// TIA Portal project "HEAT-1-CADIZ-V16" (V20) (continued)
REGION Network 5
   RUNG wire#powerrail
      "ToolChange_DB"(kukaCmdOpenCover := "kukaCmdOpenCover", kukaCmdCloseCover := "kukaCmdCloseCover", kukaCmdUnlockMps := "kukaCmdUnlockMps", kukaCmdSafeForChange := true, dockSensorToolInPosition := "dockSensorToolInPosition", dockSensorCoverClosed := "dockSensorCoverClosed", dockSensorCoverOpen := "dockSensorCoverOpen", robotSensorMpsUnlocked := "robotSensorMpsUnlocked", robotSensorMpsLocked := "robotSensorMpsLocked", robotSensorMpsCoupled := "robotSensorMpsCoupled", robotSensorMpsCtrlAirPressureOk := "robotSensorMpsCtrlAirPressureOk", resetFault :=, dockValveCoverOpenOn => "dockValveCoverOpenOn", dockValveCoverCloseOn => "dockValveCoverCloseOn", dockValveV2UnlockOn => "dockValveV2UnlockOn", kukaFeedbackDockCoverOpen => "kukaFeedbackDockCoverOpen", kukaFeedbackDockCoverClosed => "kukaFeedbackDockCoverClosed", kukaFeedbackRobotMpsUnlocked => "kukaFeedbackRobotMpsUnlocked", kukaFeedbackRobotMpsLocked => "kukaFeedbackRobotMpsLocked", kukaFeedbackRobotMpsCoupled => "kukaFeedbackRobotMpsCoupled", kukaFeedbackMpsCtrlAirPressureOk => "kukaFeedbackRobotMpsCtrlAirPressureOk", kukaFeedbackDockToolInPosition => "kukaFeedbackDockToolInPosition", diagStep =>, diagFault =>, diagFaultCode =>)
   END_RUNG
   // the same network as SCL:
   "ToolChange_DB"(kukaCmdOpenCover := "kukaCmdOpenCover",   // "ToolChange"
                   kukaCmdCloseCover := "kukaCmdCloseCover",
                   kukaCmdUnlockMps := "kukaCmdUnlockMps",
                   kukaCmdSafeForChange := true,
                   dockSensorToolInPosition := "dockSensorToolInPosition",
                   dockSensorCoverClosed := "dockSensorCoverClosed",
                   dockSensorCoverOpen := "dockSensorCoverOpen",
                   robotSensorMpsUnlocked := "robotSensorMpsUnlocked",
                   robotSensorMpsLocked := "robotSensorMpsLocked",
                   robotSensorMpsCoupled := "robotSensorMpsCoupled",
                   robotSensorMpsCtrlAirPressureOk := "robotSensorMpsCtrlAirPressureOk",
                   dockValveCoverOpenOn => "dockValveCoverOpenOn",
                   dockValveCoverCloseOn => "dockValveCoverCloseOn",
                   dockValveV2UnlockOn => "dockValveV2UnlockOn",
                   kukaFeedbackDockCoverOpen => "kukaFeedbackDockCoverOpen",
                   kukaFeedbackDockCoverClosed => "kukaFeedbackDockCoverClosed",
                   kukaFeedbackRobotMpsUnlocked => "kukaFeedbackRobotMpsUnlocked",
                   kukaFeedbackRobotMpsLocked => "kukaFeedbackRobotMpsLocked",
                   kukaFeedbackRobotMpsCoupled => "kukaFeedbackRobotMpsCoupled",
                   kukaFeedbackMpsCtrlAirPressureOk => "kukaFeedbackRobotMpsCtrlAirPressureOk",
                   kukaFeedbackDockToolInPosition => "kukaFeedbackDockToolInPosition");
END_REGION
END_FUNCTION_BLOCK

FUNCTION_BLOCK "SupervisorSeq"   // FB22, LAD
{ S7_Optimized_Access := 'TRUE' }
VERSION : 0.1
   VAR_INPUT
      T_Heartbeat : Time := T#1000ms;   // Periodo del heartbeat PLC
      T_IdCheck : Time := T#2000ms;   // Duración simulada de Identification (comprobaciones)
      enable : Bool;   // Habilita FB -> PLC.plc_ok
      QR_Ready : Bool;   // Hay un ID de carrito leído
      CarriageID : String;   // ID de carrito leído por QR
      TeachAtStart : Bool;   // Teaching (pág. 4): robot en punto de inicio de la siguiente trayectoria
      AtPerspex : Bool;   // PA check (Perspex) y Balancing (pág. 6): Robot posicionado en Perspex
      AtGainPos : Bool;   // Gain (pág. 7) -Robot posicionado para Gain
      AtTCGPos : Bool;   // TCG (pág. 8) — multiposición Robot en la posición TCG actual
      AtRefScanStart : Bool;   // Robot listo para Scan Ref
      AtInspScanStart : Bool;   // Robot listo para Scan Insp
      RefScanFinished : Bool;   // Trayectoria de referencia terminada (robot/UT)
      InspScanFinished : Bool;   // Trayectoria de inspección terminada (robot/UT)
      StartUSReady : Bool := TRUE;   // StartUS (pág. 5): end-effector y precondiciones listas -- True cuando “previous task done”
      MarkingDone : Bool;   // Pre-eval / marcado (pág. 13) -Resultado del marcado (true=OK)
      CmdStopUS : Bool;   // Orden local para Stop US
      CmdBreakUS : Bool;   // Pulso local Break US
      CmdUnbreakUS : Bool;   // Pulso local Unbreak US
   END_VAR
   VAR_OUTPUT
      ActiveStep : Int;   // Espejo local de PLC.step_plc
      AckSourceDbg : Int;   // Código de fuente de ACK (debug local)
      TCG_NextPosReq : Bool;   // PULSO 1 ciclo: mover a la SIGUIENTE posición TCG
      TCG_AdjustMode : Bool;   // LATCH: TRUE mientras estamos en “ajuste TCG”
   END_VAR
   VAR
      tHeartbeat : TON_TIME;
      tIdCheck : TON_TIME;
      hbGate : Bool;
      idCheckActive : Bool;
      prevStep : Int := -32768;
      firstScan : Bool;
      teachWasRunning : Bool;
      startUSWasRunning : Bool;
      elemWasRunning : Bool;
      balWasRunning : Bool;
      gainWasRunning : Bool;
      tcgWasInProgress : Bool;
      scanRefWasRunning : Bool;
      scanInspWasRunning : Bool;
      stopUSWasRunning : Bool;
      AckActive : Bool;   // ACK centralizado
      AckSource : Int;   // Qué petición estamos reconociendo
      evTCGNext : Bool;   // Eventos 1-ciclo que consume la máquina de estados
      evReqRefPart : Bool;
      evReqStopCycle : Bool;
      evReqTCGAdj : Bool;
      evReqVerif : Bool;
      evReqPreEval : Bool;
      evReqIdentState : Bool;
      carriageLatched : Bool;   // Otras memorias- para no reenviar ID cada ciclo
      mBreak : Bool;   // flanco Break US
      mUnbreak : Bool;   // flanco Unbreak US
      validScanParams : Bool;   // helper para scans
      waitingNextTCGPos : Bool;   // TRUE: esperar nueva posición antes de rearmar tcg_ready
   END_VAR
   VAR CONSTANT
      cSTEP_ID : Int := 1;   // // Pasos (según resumen del PDF, pág. 1)
      cSTEP_TEACH : Int := 2;
      cSTEP_STARTUS : Int := 3;
      cSTEP_PA_BAL : Int := 4;
      cSTEP_GAIN : Int := 5;
      cSTEP_TCG : Int := 6;
      cSTEP_SCAN_REF : Int := 7;
      cSTEP_SCAN_INSP : Int := 8;
      cSTEP_SCAN_REF_VERIF : Int := 9;
      cSTEP_PRE_EVAL : Int := 10;
      cACK_NONE : Int;   // // Fuentes de ACK (págs. 8, 11, 12)
      cACK_TCG_NEXT : Int := 1;
      cACK_REQ_REF : Int := 2;
      cACK_REQ_STOP : Int := 3;
      cACK_REQ_TCG_ADJ : Int := 4;
      cACK_REQ_VERIF : Int := 5;
      cACK_REQ_PRE_EVAL : Int := 6;
      cACK_REQ_IDENT_STATE : Int := 7;
   END_VAR
BEGIN

REGION Network 1 (SCL)
   // ------------------------------------------------------------------
   // 0) Servicios globales (Heartbeat, housekeeping) — vars generales (pág. 2)
   // ------------------------------------------------------------------
   "PlcStatus".plcOk := #enable;         // espejo de habilitación

   // Heartbeat PLC: toggle con TON (patrón de "compuerta")
   // hbGate se pone TRUE -> TON corre hasta PT -> tHeartbeat.Q = TRUE -> togglamos
   // y bajamos hbGate para reiniciar el ciclo.
   #tHeartbeat(IN := #hbGate,
               PT := #T_Heartbeat);
   IF NOT #hbGate THEN
       #hbGate := TRUE;
   ELSIF #tHeartbeat.Q THEN
       "PlcStatus".heartbeatPlc := NOT "PlcStatus".heartbeatPlc;
       #hbGate := FALSE;
   END_IF;

   // Normalizar paso y espejarlo a salida
   IF ("PlcStatus".stepPlc < #cSTEP_ID) OR ("PlcStatus".stepPlc > #cSTEP_PRE_EVAL) THEN
       "PlcStatus".stepPlc := #cSTEP_ID;
   END_IF;
   #ActiveStep := "PlcStatus".stepPlc;

   // firstScan: 1 ciclo al entrar en cada paso -> útil para resets seguros
   #firstScan := ("PlcStatus".stepPlc <> #prevStep);
   IF #firstScan THEN
       // Limpiamos cualquier "ready/start" que no deba arrastrarse al paso nuevo
       "PlcStatus".startUsReady := FALSE;
       "PlcStatus".stopUsReady := FALSE;
       "PlcStatus".paCheckReady := FALSE;
       "PlcStatus".gainReady := FALSE;
       "PlcStatus".tcgReady := FALSE;
       "PlcStatus".scanRefStart := FALSE;
       "PlcStatus".scanInspStart := FALSE;
       "PlcStatus".markRunning := FALSE;

       // reset de “había arrancado”
       #teachWasRunning := FALSE;
       #startUSWasRunning := FALSE;
       #elemWasRunning := FALSE;
       #balWasRunning := FALSE;
       #gainWasRunning := FALSE;
       #tcgWasInProgress := FALSE;
       #scanRefWasRunning := FALSE;
       #scanInspWasRunning := FALSE;

       // Señales generales de identificación
       "PlcStatus".idRunning := FALSE;

        //TCG: al entrar, exige confirmación de posición actual
       #waitingNextTCGPos := ("PlcStatus".stepPlc = #cSTEP_TCG) AND (NOT #AtTCGPos);
       // Salida auxiliar de ajuste TCG se limpia al cambiar de paso
       IF "PlcStatus".stepPlc <> #cSTEP_TCG THEN
           #TCG_AdjustMode := FALSE;
       END_IF;

       #prevStep := "PlcStatus".stepPlc;
   END_IF;

   // ------------------------------------------------------------------
   // [1] Gestor centralizado de ACK — TCG / Verif / PreEval / BackToID
   //     Idea: mientras una req_* esté a TRUE, PLC.acknowledge = TRUE.
   //     Cuando la req_* baja a FALSE, soltamos acknowledge y generamos
   //     un evento de 1 ciclo (evXXXX) para que el CASE tome decisiones.
   //     (ver págs. 8, 11, 12)
   // ------------------------------------------------------------------
   IF NOT #AckActive THEN
       // Tomamos la PRIMERA req_* que esté activa (prioridad de arriba a abajo)
       IF "SupervisorCmd".tcgNextStep THEN
           #AckActive := TRUE;
           #AckSource := #cACK_TCG_NEXT;
       ELSIF "SupervisorCmd".reqRefPart THEN
           #AckActive := TRUE;
           #AckSource := #cACK_REQ_REF;
       ELSIF "SupervisorCmd".reqStopCycle THEN
           #AckActive := TRUE;
           #AckSource := #cACK_REQ_STOP;
       ELSIF "SupervisorCmd".reqTcgAdj THEN
           #AckActive := TRUE;
           #AckSource := #cACK_REQ_TCG_ADJ;
       ELSIF "SupervisorCmd".reqVerif THEN
           #AckActive := TRUE;
           #AckSource := #cACK_REQ_VERIF;
       ELSIF "SupervisorCmd".reqPreEval THEN
           #AckActive := TRUE;
           #AckSource := #cACK_REQ_PRE_EVAL;
       ELSIF "SupervisorCmd".reqIdentificationState THEN
           #AckActive := TRUE;
           #AckSource := #cACK_REQ_IDENT_STATE;
       ELSE
           #AckSource := #cACK_NONE;
           #AckActive := FALSE;
       END_IF;
   END_IF;

   // Ejecutamos el reconocimiento según fuente
   CASE #AckSource OF
       #cACK_TCG_NEXT:
           "PlcStatus".acknowledge := TRUE;
           IF NOT "SupervisorCmd".tcgNextStep THEN
               // Fin del reconocimiento -> soltar y generar evento
               "PlcStatus".acknowledge := FALSE;
               #AckActive := FALSE;
               #AckSource := #cACK_NONE;
               #evTCGNext := TRUE;      // “pasar a siguiente pos” (p. 8)
           END_IF;

       #cACK_REQ_REF:
           "PlcStatus".acknowledge := TRUE;
           IF NOT "SupervisorCmd".reqRefPart THEN
               "PlcStatus".acknowledge := FALSE;
               #AckActive := FALSE;
               #AckSource := #cACK_NONE;
               #evReqRefPart := TRUE;// ir a Scan Ref (p. 8 → a)
           END_IF;

       #cACK_REQ_STOP:
           "PlcStatus".acknowledge := TRUE;
           IF NOT "SupervisorCmd".reqStopCycle THEN
               "PlcStatus".acknowledge := FALSE;
               #AckActive := FALSE;
               #AckSource := #cACK_NONE;
               #evReqStopCycle := TRUE; // cancelar ciclo (p. 8 → b)
           END_IF;

       #cACK_REQ_TCG_ADJ:
           "PlcStatus".acknowledge := TRUE;
           IF NOT "SupervisorCmd".reqTcgAdj THEN
               "PlcStatus".acknowledge := FALSE;
               #AckActive := FALSE;
               #AckSource := #cACK_NONE;
               #evReqTCGAdj := TRUE; // Seguir en TCG en modo ajuste (p. 8 → c)
           END_IF;

       #cACK_REQ_VERIF:
           "PlcStatus".acknowledge := TRUE;
           IF NOT "SupervisorCmd".reqVerif THEN
               "PlcStatus".acknowledge := FALSE;
               #AckActive := FALSE;
               #AckSource := #cACK_NONE;
               #evReqVerif := TRUE;   // Ir a verificación (p. 11)
           END_IF;

       #cACK_REQ_PRE_EVAL:
           "PlcStatus".acknowledge := TRUE;
           IF NOT "SupervisorCmd".reqPreEval THEN
               "PlcStatus".acknowledge := FALSE;
               #AckActive := FALSE;
               #AckSource := #cACK_NONE;
               #evReqPreEval := TRUE;  // Ir a Pre-eval (p. 12 → a)
           END_IF;

       #cACK_REQ_IDENT_STATE:
           "PlcStatus".acknowledge := TRUE;
           IF NOT "SupervisorCmd".reqIdentificationState THEN
               "PlcStatus".acknowledge := FALSE;
               #AckActive := FALSE;
               #AckSource := #cACK_NONE;
               #evReqIdentState := TRUE; //olver a Identification (p. 12 → b, p. 13)
           END_IF;

       ELSE
           "PlcStatus".acknowledge := FALSE;
   END_CASE;

   #AckSourceDbg := #AckSource;   // salida de diagnóstico local

   // ------------------------------------------------------------------
   // 2) MÁQUINA DE ESTADOS PRINCIPAL (CASE) — pasos del PDF
   // ------------------------------------------------------------------
   CASE "PlcStatus".stepPlc OF

           // ===============================================================
           // 1) IDENTIFICATION (pág. 3)
           // ===============================================================
       #cSTEP_ID:
           // --- Handshake de carriage ID ---
           // FÍSICO: lectura real de QR/PNs/params en HMI/Supervisor.
           // El PLC refleja ID leído y valida condiciones base (safety, agua, robot OK).
           // Supervisor.req_carriage_id = TRUE -> el PLC debe mandar:
           //   PLC.carriage_Id (string) y PLC.new_carriage_Id = TRUE
           // Mientras dure la petición. Al bajar la petición, el PLC
           // limpia new_carriage_Id y deja de enviar.
           // req_carriage_id: enviar ID nuevo UNA VEZ mientras Supervisor lo solicite
           IF "SupervisorCmd".reqCarriageId THEN
               IF #QR_Ready AND NOT #carriageLatched THEN
                   "PlcStatus".carriageId := #CarriageID; // escribimos el ID leído
                   "PlcStatus".newCarriageId := TRUE;     // “ID listo”
                   #carriageLatched := TRUE;              // evita rearmar en el mismo pulso
               END_IF;
           ELSE
               // fin del handshake
               "PlcStatus".newCarriageId := FALSE;
               #carriageLatched := FALSE;
           END_IF;

           // --- req_id -> identificación en curso ---
           // Cuando Supervisor pone req_id, el PLC indica id_running y,
           // tras un tiempo T_IdCheck, fija id_ok según condiciones globales.
           IF "SupervisorCmd".reqId AND NOT #idCheckActive THEN
               #idCheckActive := TRUE;
               "PlcStatus".idRunning := TRUE;
               "PlcStatus".idOk := FALSE;
               #tIdCheck(IN := TRUE,
                         PT := #T_IdCheck);  // arranca temporizador
           END_IF;

           IF #idCheckActive THEN
               #tIdCheck(IN := TRUE,
                         PT := #T_IdCheck);
               IF #tIdCheck.Q THEN
                   // Condiciones base (p. 2): enclavamientos / servicios / robot listo
                   "PlcStatus".idOk := ("PlcStatus".plcOk AND "SupervisorCmd".supervisorOk AND "PlcStatus".robotOk AND "PlcStatus".safetyOk
                   AND "PlcStatus".airOk AND "PlcStatus".inspWaterOk AND "PlcStatus".tankWaterOk);
                   "PlcStatus".idRunning := FALSE;
                   #idCheckActive := FALSE;
                   #tIdCheck(IN := FALSE,
                             PT := #T_IdCheck);

                   // Saltos según resultado y teach_req (pág. 3)
                   IF NOT "PlcStatus".idOk THEN
                       "PlcStatus".stepPlc := #cSTEP_ID; // cancelar ciclo / quedarse en identificación
                   ELSE
                       // Siguiente paso según teach_req (pág. 3)
                       IF "SupervisorCmd".teachReq THEN
                           "PlcStatus".stepPlc := #cSTEP_TEACH;
                       ELSE
                           "PlcStatus".stepPlc := #cSTEP_STARTUS;
                       END_IF;
                   END_IF;
               END_IF;
           ELSE
               // Aseguramos TON parado fuera del ciclo activo
               #tIdCheck(IN := FALSE,
                         PT := #T_IdCheck);
           END_IF;


           // ===============================================================
           // 2) TEACHING (pág. 4) — multi-PN: rearmar teach_ready por PN
           // FÍSICO: si la herramienta necesaria para teaching no está montada,
           // el KUKA cambia en Staübli al stand indicado (usa Supervisor.end-effector).
           // Luego, el KUKA se mueve al INICIO del PN siguiente y pone un bit de “en posición”.
           // Ese bit alimenta TeachAtStart=TRUE. Entonces EL PLC arma teach_ready (p. 4).
           // Repetir por cada PN mientras teach_app_running=TRUE.
           // ===============================================================
           (*  #cSTEP_TEACH:

            // Mientras la app de teaching esté abierta, debemos rearmar teach_ready
            // cada vez que el robot esté en el inicio del siguiente PN (TeachAtStart).
           IF "SupervisorCmd".teachAppRunning THEN
               // "Listo para enseñar" SOLO si NO está corriendo y robot en inicio PN              
               IF (NOT Supervisor.teach_running) AND #TeachAtStart THEN
                   "PlcStatus".teach_ready := TRUE; // // el láser/soft podrá iniciar teaching
               END_IF;

             // Al arrancar trayectoria de teaching -> soltamos ready
               IF Supervisor.teach_running THEN
                   PLC.teach_ready := FALSE;
                   #teachWasRunning := TRUE; // marcamos que empezó realmente
               END_IF;

                  // Al terminar una trayectoria (teach_running pasa a FALSE)
               IF (NOT Supervisor.teach_running) AND #teachWasRunning THEN
                   #teachWasRunning := FALSE; // fin de una trayectoria teaching
                    // Si siguen más PNs, se rearmará arriba (TeachAtStart=TRUE).
               END_IF;
           ELSE
                // Cierre de la app -> decidimos salto en base a teach_state (pág. 4)
               IF Supervisor.teach_state THEN
                   PLC.step_plc := #cSTEP_STARTUS;
               ELSE
                   PLC.step_plc := #cSTEP_ID;
               END_IF;
           END_IF;*)




           // ===============================================================
           // 3) START US (pág. 5) — armar cuando “previous task done”
           // FÍSICO: KUKA AUT EXT cambia (si hace falta) al efector de INSPECCIÓN
           // requerido (Supervisor.end-effector, p. 1). Cuando:
           //   - Herramienta correcta acoplada (Staübli OK),
           //   - servicios/enclavamientos OK (safety/air/water/tank),
           //   - robot en posición segura para inicializar el UT,
           // tu secuenciador pone StartUSReady=TRUE. El PLC arma start_us_ready.
           // Supervisor hace init UT (start_us_running/state_us). (p. 5)
           // ===============================================================
       #cSTEP_STARTUS:

           // Solo armamos start_us_ready si “previous task done” (StartUSReady)
           // y el Supervisor aún no ha arrancado.
           IF #StartUSReady AND NOT "SupervisorCmd".startUsRunning THEN
               "PlcStatus".startUsReady := TRUE; // → Supervisor puede iniciar
           END_IF;

           // Al comenzar la inicialización, soltamos el ready
           IF "SupervisorCmd".startUsRunning THEN
               "PlcStatus".startUsReady := FALSE;
               #startUSWasRunning := TRUE;
           END_IF;

           // Al finalizar la inicialización, Supervisor deja de correr y publica state_us
           IF (NOT "SupervisorCmd".startUsRunning) AND #startUSWasRunning THEN
               #startUSWasRunning := FALSE;
               IF NOT "SupervisorCmd".stateUs THEN
                   "PlcStatus".stepPlc := #cSTEP_ID; // fallo init US -> cancelar
               ELSE
                   IF "SupervisorCmd".paCheckReq THEN
                       "PlcStatus".stepPlc := #cSTEP_PA_BAL; // a) ir a PA-check (p. 5)
                   ELSE
                       "PlcStatus".stepPlc := #cSTEP_GAIN;   // b) ir a Gain (p. 5)
                   END_IF;
               END_IF;
           END_IF;

           // ===============================================================
           // 4) DEAD ELEMENT CHECK & BALANCING (pág. 6)
           //FÍSICO: KUKA va a la pieza Perspex de calibración y, cuando está en
           // posición estática, tu lógica pone AtPerspex=TRUE. El PLC arma
           // pa_check_ready y el Supervisor ejecuta elem_running/bal_running (p. 6).
           // ===============================================================
       #cSTEP_PA_BAL:

           // Dead elements en Perspex: el PLC pone pa_check_ready SOLO si
           // el robot ya está en la pieza Perspex y aún no corre elem_running
           IF #AtPerspex AND NOT "SupervisorCmd".elemRunning THEN
               "PlcStatus".paCheckReady := TRUE;
           END_IF;

           // Al iniciar la comprobación de dead elements soltamos ready
           IF "SupervisorCmd".elemRunning THEN
               "PlcStatus".paCheckReady := FALSE;
               #elemWasRunning := TRUE;
           END_IF;

           // Fin de dead elements -> miramos elem_state y encadenamos Balancing
           IF (NOT "SupervisorCmd".elemRunning) AND #elemWasRunning THEN
               #elemWasRunning := FALSE;
               IF NOT "SupervisorCmd".elemState THEN
                   "PlcStatus".stepPlc := #cSTEP_ID;
               ELSE
                   // Cascada a balancing (misma posición Perspex) (p. 6)
                   IF "SupervisorCmd".balRunning THEN
                       #balWasRunning := TRUE;
                   END_IF;

                   IF (NOT "SupervisorCmd".balRunning) AND #balWasRunning THEN
                       #balWasRunning := FALSE;
                       IF "SupervisorCmd".balState THEN
                           "PlcStatus".stepPlc := #cSTEP_GAIN;
                       ELSE
                           "PlcStatus".stepPlc := #cSTEP_ID;
                       END_IF;
                   END_IF;
               END_IF;
           END_IF;

           // ===============================================================
           // 5) GAIN ADJUSTMENT (pág. 7)
           // FÍSICO: KUKA se posiciona en la referencia para ganancia estática;
           // cuando está “en posición”, AtGainPos=TRUE. PLC arma gain_ready;
           // Supervisor ejecuta gain_running/gain_state y decide si ir a TCG (p. 7).
           // ===============================================================
       #cSTEP_GAIN:

           // Armamos gain_ready únicamente cuando el robot está en la posición
           // de ganancia y el supervisor todavía no corre la rutina de gain
           IF #AtGainPos AND NOT "SupervisorCmd".gainRunning THEN
               "PlcStatus".gainReady := TRUE;  // → Supervisor puede iniciar
           END_IF;

           IF "SupervisorCmd".gainRunning THEN
               "PlcStatus".gainReady := FALSE;
               #gainWasRunning := TRUE;
           END_IF;

           // Al terminar gain, ver resultado y decidir: TCG o Scan Ref
           IF (NOT "SupervisorCmd".gainRunning) AND #gainWasRunning THEN
               #gainWasRunning := FALSE;
               IF NOT "SupervisorCmd".gainState THEN
                   "PlcStatus".stepPlc := #cSTEP_ID;
               ELSE
                   IF "SupervisorCmd".tcgReq THEN
                       "PlcStatus".stepPlc := #cSTEP_TCG;
                   ELSE
                       "PlcStatus".stepPlc := #cSTEP_SCAN_REF;
                   END_IF;
               END_IF;
           END_IF;

           // ===============================================================
           // (6) TCG CHECK / ADJUSTMENT — pág. 8 (multiposición)
           // FÍSICO: KUKA recorre varias posiciones TCG. Para cada posición:
           //   - Cuando el robot está en la POSICIÓN TCG ACTUAL (estático),
           //     tu lógica pone AtTCGPos=TRUE → PLC arma tcg_ready (p. 8).
           //   - Supervisor pone tcg_in_progress=TRUE mientras mide.
           //   - Al pulsar “Next” en Supervisor (tcg_next_step=TRUE), el ACK manager
           //     emite TCG_NextPosReq (pulso) para que MUEVAS el robot a la SIGUIENTE
           //     posición; el FB bloquea el rearme (waitingNextTCGPos=TRUE) hasta que
           //     AtTCGPos vuelva a TRUE en la nueva posición (antirrebote).
           //   - Final: según req_ref_part / req_stop_cycle / req_tcg_adj (p. 8).
           // ===============================================================
       #cSTEP_TCG:

           // Confirmación de nueva posición alcanzada
           IF #waitingNextTCGPos AND #AtTCGPos THEN
               #waitingNextTCGPos := FALSE;     // nueva pos OK → se podrá rearmar ready
           END_IF;

           // Armado defensivo: tcg_ready SOLO si no hay progreso y no esperamos pos
           IF (NOT "SupervisorCmd".tcgInProgress) AND (NOT #waitingNextTCGPos) THEN
               "PlcStatus".tcgReady := TRUE;          // listo para medir en esta pos (p. 8)
           END_IF;

           IF "SupervisorCmd".tcgInProgress THEN
               "PlcStatus".tcgReady := FALSE;
               #tcgWasInProgress := TRUE;
           END_IF;

           // “Next” → mueve a la SIGUIENTE pos (tu secuenciador KUKA)
           IF #evTCGNext THEN
               #TCG_NextPosReq := TRUE;      // pulso 1 ciclo hacia tu lógica
               #waitingNextTCGPos := TRUE;      // bloquea ready hasta nueva posición
           END_IF;

           // “Ajuste TCG”
           IF #evReqTCGAdj THEN
               #TCG_AdjustMode := TRUE;        // permanecer en step 6 hasta validar
           END_IF;

           // Validación de TCG
           IF #evReqRefPart THEN
               #TCG_AdjustMode := FALSE;
               "PlcStatus".stepPlc := #cSTEP_SCAN_REF; // TCG OK → Scan Ref (p. 8)
           ELSIF #evReqStopCycle THEN
               #TCG_AdjustMode := FALSE;
               "PlcStatus".stepPlc := #cSTEP_ID;       // cancelar (p. 8)
           END_IF;



           // ===============================================================
           // (7) SCAN REFERENCE ACQUISITION — pág. 10
           // FÍSICO: KUKA carga PN/frame y se coloca en el punto de INICIO de
           // la trayectoria de referencia. Tu lógica pone AtRefScanStart=TRUE cuando
           // está en posición. El PLC solo arma scan_ref_start si además los
           // parámetros mínimos (id_scan, x_size, y_size) están válidos (p. 10).
           // ===============================================================
       #cSTEP_SCAN_REF:

           // Validación mínima de parámetros: hay PN/Frame y tamaños > 0.
           // (El PDF indica que el PLC envía id_scan, point_origin, x_size, y_size).
           #validScanParams := (LEN("PlcStatus".idScan) > 0) AND ("PlcStatus".xSize > 0.0) AND ("PlcStatus".ySize > 0.0);

           // "Robot ready" solo si parámetros OK, robot en inicio y aún no corre
           IF #AtRefScanStart AND #validScanParams AND NOT "SupervisorCmd".scanRefRunning THEN
               "PlcStatus".scanRefStart := TRUE;     // Supervisor cargará/validará y pondrá scan_ref_running
           END_IF;

           // En ejecución: opcionalmente bajar start al terminar la trayectoria
           IF "SupervisorCmd".scanRefRunning THEN
               #scanRefWasRunning := TRUE;
               IF #RefScanFinished THEN
                   "PlcStatus".scanRefStart := FALSE; // indica “fin de movimiento -> guardar”
               END_IF;
           END_IF;

           // Al terminar guardado, Supervisor baja running y publica scan_ref_state
           IF (NOT "SupervisorCmd".scanRefRunning) AND #scanRefWasRunning THEN
               #scanRefWasRunning := FALSE;
               "PlcStatus".scanRefStart := FALSE;
               IF NOT "SupervisorCmd".scanRefState THEN
                   "PlcStatus".stepPlc := #cSTEP_ID;   // error durante ref -> cancelar
               ELSE
                   "PlcStatus".stepPlc := #cSTEP_SCAN_INSP;
               END_IF;
           END_IF;

           // ===============================================================
           // (8) SCAN INSPECTION — pág. 11
           // FÍSICO: KUKA se coloca en INICIO de la(s) trayectoria(s) de inspección
           // (AtInspScanStart=TRUE). El PLC arma scan_insp_start solo si parámetros
           // válidos. Supervisor corre/guarda y luego pide verificación (req_verif) (p. 11).
           // ===============================================================
       #cSTEP_SCAN_INSP:

           // Validación mínima de parámetros: hay PN/Frame y tamaños > 0.
           // (El PDF indica que el PLC envía id_scan, point_origin, x_size, y_size).
           #validScanParams := (LEN("PlcStatus".idScan) > 0) AND ("PlcStatus".xSize > 0.0) AND ("PlcStatus".ySize > 0.0);

           // "Robot ready" solo si parámetros OK, robot en inicio y aún no corre
           IF #AtInspScanStart AND #validScanParams AND NOT "SupervisorCmd".scanInsprunning THEN
               "PlcStatus".scanInspStart := TRUE;    // Supervisor cargará y arrancará
           END_IF;

           // En ejecución: opcionalmente bajar start al terminar la trayectoria
           IF "SupervisorCmd".scanInsprunning THEN
               #scanInspWasRunning := TRUE;
               IF #InspScanFinished THEN
                   "PlcStatus".scanInspStart := FALSE; // fin de movimiento -> guardar
               END_IF;
           END_IF;

           // Al terminar guardado, Supervisor baja running y publica scan_ref_state
           IF (NOT "SupervisorCmd".scanInsprunning) AND #scanInspWasRunning THEN
               #scanInspWasRunning := FALSE;
               "PlcStatus".scanInspStart := FALSE;

               IF NOT "SupervisorCmd".scanInspState THEN
                   "PlcStatus".stepPlc := #cSTEP_ID;   // error -> cancelar
               ELSE
                   // Ir a verificación cuando el ACK manager confirme req_verif
                   IF #evReqVerif THEN
                       "PlcStatus".stepPlc := #cSTEP_SCAN_REF_VERIF;
                   END_IF;
               END_IF;
           END_IF;


           // ===============================================================
           // (9) SCAN REFERENCE VERIFICATION — pág. 12
           // FÍSICO: KUKA vuelve al INICIO de la trayectoria de verificación de ref.
           // (AtRefScanStart=TRUE). Igual patrón de parámetros/ready/running/state (p. 12).
           // Fin: Supervisor decide Pre‑eval (req_pre_eval) o nuevo ciclo (req_identification_state).
           // ===============================================================
       #cSTEP_SCAN_REF_VERIF:

           #validScanParams := (LEN("PlcStatus".idScan) > 0) AND ("PlcStatus".xSize > 0.0) AND ("PlcStatus".ySize > 0.0);

           IF #AtRefScanStart AND #validScanParams AND NOT "SupervisorCmd".scanRefRunning THEN
               "PlcStatus".scanRefStart := TRUE;     // Robot listo para verificación de ref
           END_IF;

           IF "SupervisorCmd".scanRefRunning THEN
               #scanRefWasRunning := TRUE;
           END_IF;

           IF (NOT "SupervisorCmd".scanRefRunning) AND #scanRefWasRunning THEN
               #scanRefWasRunning := FALSE;
               "PlcStatus".scanRefStart := FALSE;

               IF NOT "SupervisorCmd".scanRefState THEN
                   "PlcStatus".stepPlc := #cSTEP_ID;
               ELSE
                   // a) Pre‑eval   b) Volver a Identification
                   IF #evReqPreEval THEN
                       "PlcStatus".stepPlc := #cSTEP_PRE_EVAL;
                   ELSIF #evReqIdentState THEN
                       "PlcStatus".stepPlc := #cSTEP_ID;
                   END_IF;
               END_IF;
           END_IF;

           // ===============================================================
           // (10) PRE‑EVALUATION / MARKING — pág. 13
           // FÍSICO: si la herramienta de marcado no está montada, el KUKA cambia
           // en Staübli al stand de “marking” según requiera el proceso; tras estar
           // listo se puede marcar (Supervisor.req_mark). El resultado físico del
           // marcado tu lógica lo refleja en MarkingDone=TRUE/FALSE (p. 13).
           // También se puede arrancar un nuevo ciclo (req_identification_state).
           // ===============================================================
       #cSTEP_PRE_EVAL:

           // b) Volver a inicio (nuevo ciclo)
           IF #evReqIdentState THEN
               "PlcStatus".stepPlc := #cSTEP_ID;
           END_IF;

           // a) Marcado: si Supervisor.req_mark, ejecutamos el ciclo simple:
           //   - mark_running TRUE durante la acción
           //   - mark_state según resultado físico (MarkingDone)
           IF "SupervisorCmd".reqMark THEN
               "PlcStatus".markState := FALSE;      // reset explícito del estado
               "PlcStatus".markRunning := TRUE;       // marcando...

               "PlcStatus".markState := #MarkingDone; // resultado del efector externo

               "PlcStatus".markRunning := FALSE;      // fin de marcado (Supervisor bajará req_mark)
           END_IF;


           // Fallback de seguridad
       ELSE
           "PlcStatus".stepPlc := #cSTEP_ID;


   END_CASE;


   // ------------------------------------------------------------------
   // [3] Servicios FUERA DE CICLO — StopUS / Rescanning / Break&Unbreak / Error
   // ------------------------------------------------------------------

   // Stop US (pág. 9). El PLC puede lanzar stop_us_ready cuando proceda
   // (por ejemplo, antes de cambiar efector con el agua aún presente).
   IF #CmdStopUS THEN
       "PlcStatus".stopUsReady := TRUE;
   END_IF;

   // Handshake de StopUS: Supervisor pone stop_us_running mientras ejecuta;
   // cuando termina, bajará stop_us_running y aquí soltamos stop_us_ready.
   IF "PlcStatus".stopUsReady THEN
       IF "SupervisorCmd".stopUsRunning THEN
           #stopUSWasRunning := TRUE;
       END_IF;

       IF (NOT "SupervisorCmd".stopUsRunning) AND #stopUSWasRunning THEN
           #stopUSWasRunning := FALSE;
           "PlcStatus".stopUsReady := FALSE; // handshake completado
       END_IF;
   ELSE
       #stopUSWasRunning := FALSE;
   END_IF;

   // Break / Unbreak (pág. 14): pulsos de 1 ciclo a petición local
   IF (#CmdBreakUS AND NOT #mBreak) THEN
       "PlcStatus".breakUs := TRUE;   // Supervisor cambiará state_us en consecuencia
   ELSE
       "PlcStatus".breakUs := FALSE;
   END_IF;
   #mBreak := #CmdBreakUS;

   IF (#CmdUnbreakUS AND NOT #mUnbreak) THEN
       "PlcStatus".unbreakUs := TRUE; // Supervisor volverá a poner state_us TRUE
   ELSE
       "PlcStatus".unbreakUs := FALSE;
   END_IF;
   #mUnbreak := #CmdUnbreakUS;

   // Rescanning (pág. 15): reflejar que el robot está listo para rebobinar
   IF "SupervisorCmd".rescanning THEN
       "PlcStatus".robotRescanning := TRUE;
   ELSE
       "PlcStatus".robotRescanning := FALSE;
   END_IF;

   // Gestión de errores (pág. 16): mantener acknowledge_error en TRUE
   // mientras dure error_occured; soltar cuando se limpie.
   IF "SupervisorCmd".errorOcurred THEN
       "PlcStatus".acknowledgeError := TRUE;
   ELSE
       "PlcStatus".acknowledgeError := FALSE;
   END_IF;

   // ---- Limpieza de eventos de 1 ciclo (siempre al final del scan) ----
   #evTCGNext := FALSE;
   #evReqRefPart := FALSE;
   #evReqStopCycle := FALSE;
   #evReqTCGAdj := FALSE;
   #evReqVerif := FALSE;
   #evReqPreEval := FALSE;
   #evReqIdentState := FALSE;
END_REGION
END_FUNCTION_BLOCK

ORGANIZATION_BLOCK "Main"   // OB1, LAD, ProgramCycle
TITLE = "Main Program Sweep (Cycle)"
{ S7_Optimized_Access := 'TRUE' }
VERSION : 0.1
   VAR_INPUT
      Initial_Call : Bool;   // Initial call of this OB
      Remanence : Bool;   // =True, if remanent data are available
   END_VAR
   VAR_TEMP
      evtEnterSrv : Bool;   // // Eventos de modo service jog
      evtEnterAuto : Bool;   // // Eventos de modo auto
      muxSelStb : Bool;
      muxStartStb : Bool;
      muxPgno : Byte;
      u : UDInt;
   END_VAR
BEGIN

REGION Network 1 (SCL): // ====================== READ (%I) ======================
   // // —— Enlaza estos símbolos a tus %I en el árbol de dispositivos ——
   //   // EStop_DI, SafeDoor_DI, AirPressure_DI, WaterInsp_DI, WaterTank_DI, RobotReady_DI, ...
END_REGION

REGION Network 2: // 1) Árbitro de modo: decide y emite
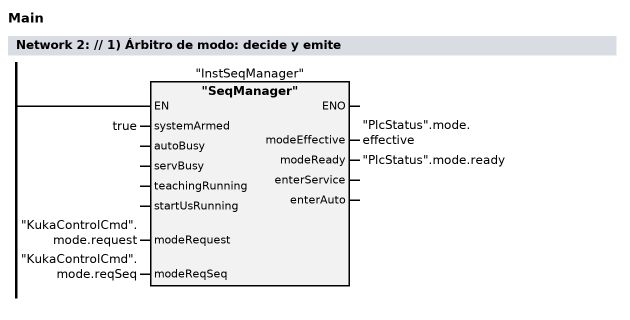
   RUNG wire#powerrail
      "InstSeqManager"(systemArmed := true, autoBusy :=, servBusy :=, teachingRunning :=, startUsRunning :=, modeRequest := "KukaControlCmd".mode.request, modeReqSeq := "KukaControlCmd".mode.reqSeq, modeEffective => "PlcStatus".mode.effective, modeReady => "PlcStatus".mode.ready, enterService =>, enterAuto =>)
   END_RUNG
   // the same network as SCL:
   "InstSeqManager"(systemArmed := true,   // "SeqManager"
                    modeRequest := "KukaControlCmd".mode.request,
                    modeReqSeq := "KukaControlCmd".mode.reqSeq,
                    modeEffective => "PlcStatus".mode.effective,
                    modeReady => "PlcStatus".mode.ready);
END_REGION

REGION Network 3 (SCL): // 2) Ejecuta o service o Auto
       IF "PlcStatus".mode.effective = 1 THEN
           // SUPERVISOR : Mode Effective = 1
           "InstSupervisorSeq"();
       ELSE
           // KUKACONTROL: Mode Effective = 0
           "InstKukaControlSeq"();
       END_IF;
END_REGION
END_ORGANIZATION_BLOCK

// folder: 10. System/Utilities

FUNCTION_BLOCK "ClockPulse"   // FB67, LAD
{ S7_Optimized_Access := 'TRUE' }
VERSION : 0.1
BEGIN
END_FUNCTION_BLOCK

// folder: 20. Robot Services/AutoExt

FUNCTION_BLOCK "AutoExtSeq"   // FB31, LAD
{ S7_Optimized_Access := 'TRUE' }
VERSION : 0.1
   VAR_INPUT
      enable : Bool;   // // habilita interfaz
      startCmd : Bool;   // // flanco de arranque
      ProgramNo : Byte;   // / nº CASE (1..255)
      AutoAck : Bool;   // // auto-confirmar STOPMESS
   END_VAR
   VAR
      rStart : R_TRIG;
      Static_1 : Bool;
      fReq : F_TRIG;
      pending : Bool;   // // hay pedido en curso
      running : Bool;   // // PRO_ACT latcheado
      pgnoLat : Byte;   // // PGNO latcheado
      tpStart : TP_TIME;
      tpAck : TP_TIME;
      rStop : R_TRIG;
   END_VAR
BEGIN

REGION Network 2 (SCL): // ---- detectar solicitud de arranque ----
END_REGION

REGION Network 3 (SCL): Paridad
END_REGION

REGION Network 4 (SCL): // ---- VALID solo mientras PGNO_REQ=1 y hay pedido ----
END_REGION

REGION Network 5 (SCL): // ---- cuando PGNO_REQ baja -> pulso de EXT_START ---
END_REGION

REGION Network 6 (SCL): // ---- auto-confirmar mensajes cuando aparezcan ----
END_REGION

REGION Network 7 (SCL): ---- seguimiento de ejecución y liberación de 'pending' ----
END_REGION
END_FUNCTION_BLOCK

// folder: 20. Robot Services/Mov Manual

FUNCTION_BLOCK "TcpJogging"   // FB5, LAD
{ S7_Optimized_Access := 'TRUE' }
VERSION : 0.1
   VAR_INPUT
      "buttonX+" : Bool;
      "buttonX-" : Bool;
      "buttonY+" : Bool;
      "buttonY-" : Bool;
      "buttonZ+" : Bool;
      "buttonZ-" : Bool;
      "buttonE1+" : Bool;
      "buttonE1-" : Bool;
   END_VAR
BEGIN

REGION Network 1 (SCL): Mapea los valores de los botones de WF
   IF "PlcStatus".mode.effective = 0 THEN

       "Tag_1" := TRUE;
       //MOV X,Y,Z
       //%Q630.0 = buttonX+
       //%Q630.1 = buttonX-
       //%Q630.2 = buttonY+
       //%Q630.3 = buttonY-
       //%Q630.4 = buttonZ+
       //%Q630.5 = buttonZ-
       //MOV A,B,C
       //%Q630.6 = buttonWF +A
       //%Q630.7 = buttonWF -A
       //%Q631.0 = buttonWF +B
       //%Q631.1 = buttonWF -B
       //%Q631.2 = buttonWF +C
       //%Q631.3 = buttonWF -C
       //Mov E1
       //%Q631.4 = buttonWF +E1
       //%Q631.5 = buttonWF -E1

   ELSE
       //%Q631.1 = buttonWF -B
       "Tag_1" := FALSE;
   END_IF;
END_REGION
END_FUNCTION_BLOCK

FUNCTION_BLOCK "TcpTarget"   // FB11, LAD
{ S7_Optimized_Access := 'TRUE' }
VERSION : 0.1
   VAR_INPUT
      KukaControlCmdCode : UInt;
      KukaControlCmdSeq : UInt;
      KukaControlCmdProfileRequestId : UInt;
      KukaControlCmdToolRequestId : UInt;
      KukaControlCmdBaseRequestId : UInt;
      KukaControlCmdProgramRequestId : UInt;
      KukaControlTcpTargetX_mm : LReal;
      KukaControlTcpTargetY_mm : LReal;
      KukaControlTcpTargetZ_mm : LReal;
      kukaControlE1Target_mm : LReal;
      KukaControlCmdCancelGo : Bool;
      KukaControlCmdPauseGo : Bool;
      KukaControlCmdResumeGo : Bool;
   END_VAR
   VAR_OUTPUT
      moveCodeKuka : Word;
      profileReqId : Word;
      baseReqId : Word;
      toolReqId : Word;
      programReqId : Word;
      x_mmHe : DWord;
      y_mmHe : DWord;
      z_mmHe : DWord;
      e_mmHe : DWord;
      PlcStatusExecDone : Bool;
      PlcStatusExecAccepted : Bool;
      PlcStatusExecAckSeq : UInt;
      PlcStatusExecBusy : Bool;
      PlcStatusExecError : Bool;
      PlcStatusExecErrorCode : DWord;
      PlcStatusExecLastCode : UInt;
      PlcStatusCancelAck : Bool;
      PlcStatusPauseAck : Bool;
      PlcStatusResumeAck : Bool;
      PlcStatusExecPaused : Bool;
   END_VAR
   VAR
      lastSeq : UInt;
      lastCode : UInt;
      state : Int;
      tmoMove : TON_TIME;
      rbDoneEdge : R_TRIG;
      _cancelInFlight : Bool := false;   // marca que el DONE que venga es por cancelación
      _isMotion : Bool;   // helper para saber si el code es de movimiento
   END_VAR
   VAR_TEMP
      x_dint : DInt;
      y_dint : DInt;
      z_dint : DInt;
      n_dint : DInt;
      code_int : UInt;
      tool_int : UInt;
   END_VAR
BEGIN

REGION Network 1 (SCL)
   // =================== Canal asíncrono ExecCtrl ====================
   // Handshake por nivel: <Go> de HMI -> PLC -> KRC, y cierre al recibir <Ack> del KRC.
   // Al cerrar, reflejamos el Ack hacia HMI y actualizamos PlcStatusExecPaused.

   // ---- CANCEL ----
   IF (#KukaControlCmdCancelGo <> #PlcStatusCancelAck) THEN
       "cancelGo" := #KukaControlCmdCancelGo;   // propaga al KRC
       #_cancelInFlight := TRUE;              // esperamos DONE por cancel
       // cerrar cuando el KRC confirme
       IF ("cancelAck" = "cancelGo") THEN
           #PlcStatusCancelAck := #KukaControlCmdCancelGo;  // cierra HMI
           #PlcStatusExecPaused := FALSE;                 // cancel limpia pausa (si la había)
       END_IF;
   END_IF;

   // ---- PAUSE ----
   IF (#KukaControlCmdPauseGo <> #PlcStatusPauseAck) THEN
       "pauseGo" := #KukaControlCmdPauseGo;     // propaga al KRC
       IF ("pauseAck" = "pauseGo") THEN
           #PlcStatusPauseAck := #KukaControlCmdPauseGo;    // cierra HMI
           #PlcStatusExecPaused := TRUE;                   // queda en pausa reanudable
       END_IF;
   END_IF;

   // ---- RESUME ----
   IF (#KukaControlCmdResumeGo <> #PlcStatusResumeAck) THEN
       "resumeGo" := #KukaControlCmdResumeGo;   // propaga al KRC
       IF ("resumeAck" = "resumeGo") THEN
           #PlcStatusResumeAck := #KukaControlCmdResumeGo;  // cierra HMI
           #PlcStatusExecPaused := FALSE;                 // fuera de pausa
       END_IF;
   END_IF;

   CASE #state OF
       0: // IDLE -> GO == ACK
           #PlcStatusExecAccepted := FALSE;
           #PlcStatusExecBusy := FALSE;
           #PlcStatusExecError := FALSE;
           //#PlcStatusExecDone := FALSE;

           // Nuevo comando si llega seq distinto y hay código válido
           IF (#KukaControlCmdSeq <> #lastSeq)  THEN

               // (1) Latch del código para decidir si es movimiento
               #code_int := #KukaControlCmdCode;
               #_isMotion := (#code_int = 101) OR (#code_int = 102) OR (#code_int = 103) OR
               (#code_int = 130) OR (#code_int = 402);

               // (2) Solo disparamos si el canal está libre
               IF ("goTrigger" ="rbDone") THEN
                   // 1) Volcar dataset PNIO (tool/base/vel/target...) hacia el robot
                   // Prepara dataset hacia KUKA

                   // (opcional) bloquear nuevos movimientos si estamos en pausa
                   IF NOT (#PlcStatusExecPaused AND #_isMotion) THEN


                   //  Primero: Escalar mm → entero (µm). Ajusta el redondeo si lo prefieres TRUNC, FLOOR, etc.
                   #code_int := #KukaControlCmdCode;
                   #tool_int := #KukaControlCmdToolRequestId;
                   // 1) Usa el code local (sin swap) para decidir

                   IF #code_int = 130 THEN
                       //  Primero: Escalar mm → entero (µm). Ajusta el redondeo si lo prefieres TRUNC, FLOOR, etc.
                       #n_dint := LREAL_TO_DINT(ROUND(#kukaControlE1Target_mm));
                       // Segundo Convertir a DWORD y hacer SWAP para que el KRC lo lea correctamente
                       #e_mmHe := SWAP(DINT_TO_DWORD(#n_dint));
                   END_IF;

                   IF #code_int = 101 THEN
                       //  Primero: Escalar mm → entero (µm). Ajusta el redondeo si lo prefieres TRUNC, FLOOR, etc.
                       #x_dint := LREAL_TO_DINT(ROUND(#KukaControlTcpTargetX_mm));
                       // Segundo Convertir a DWORD y hacer SWAP para que el KRC lo lea correctamente
                       #x_mmHe := SWAP(DINT_TO_DWORD(#x_dint));
                   END_IF;

                   IF #code_int = 102 THEN
                       //  Primero: Escalar mm → entero (µm). Ajusta el redondeo si lo prefieres TRUNC, FLOOR, etc.
                       #y_dint := LREAL_TO_DINT(ROUND(#KukaControlTcpTargetY_mm));
                       // Segundo Convertir a DWORD y hacer SWAP para que el KRC lo lea correctamente
                       #y_mmHe := SWAP(DINT_TO_DWORD(#y_dint));
                   END_IF;

                   IF #code_int = 103 THEN
                       //  Primero: Escalar mm → entero (µm). Ajusta el redondeo si lo prefieres TRUNC, FLOOR, etc.
                       #z_dint := LREAL_TO_DINT(ROUND(#KukaControlTcpTargetZ_mm));
                       // Segundo Convertir a DWORD y hacer SWAP para que el KRC lo lea correctamente
                       #z_mmHe := SWAP(DINT_TO_DWORD(#z_dint));
                   END_IF;

                   IF #code_int = 201 THEN
                       // id de herramienta → WORD+SWAP
                       #toolReqId := SWAP(UINT_TO_WORD(#KukaControlCmdToolRequestId));

                   END_IF;

                   IF #code_int = 202 THEN

                       // id de herramienta → WORD+SWAP
                       #baseReqId := SWAP(UINT_TO_WORD(#KukaControlCmdBaseRequestId));

                   END_IF;

                   IF #code_int = 203 THEN

                       // id de herramienta → WORD+SWAP
                       #profileReqId := SWAP(UINT_TO_WORD(#KukaControlCmdProfileRequestId));

                   END_IF;

                   // ---------- TEACHING ----------
                   IF #code_int = 301 THEN // Teach Request
                       #programReqId := SWAP(UINT_TO_WORD(#KukaControlCmdProgramRequestId));

                   END_IF;


                   IF #code_int = 311 OR #code_int = 312 OR #code_int = 313 THEN

                       // sin parámetros adicionales
                       #programReqId := SWAP(UINT_TO_WORD(#KukaControlCmdProgramRequestId));
                   END_IF;

                   // ---------- SCAN ----------
                   IF #code_int = 401 OR #code_int = 402 THEN

                       #programReqId := SWAP(UINT_TO_WORD(#KukaControlCmdProgramRequestId)); 
                       // (opcional) velocidad por PNIO:
                       //vel_mmsHe := SWAP(#KukaControlCmd_vel_mms);          // WORD con SWAP si tu PNIO lo requiere
                       // index: mm -> µm -> DWORD + SWAP
                       //#n_dint := LREAL_TO_DINT(ROUND(#KukaControlCmd_index_mm * 1000.0));
                       //index_umHe := SWAP(DINT_TO_DWORD(#n_dint));
                   END_IF;



                   // Segundo Convertir a DWORD y hacer SWAP para que el KRC lo lea correctamente
                   #moveCodeKuka := SWAP(UINT_TO_WORD(#code_int));
                  // "moveCodeKuka" := SWAP(UINT_TO_WORD(#code_int));

                   // Dispara GO (flanco por nivel)
                   "goTrigger" := NOT "goTrigger";     // Dispara pedido

                   // Marca estado/ack interno
                   #PlcStatusExecAccepted := TRUE;
                   #PlcStatusExecBusy := TRUE;
                   #PlcStatusExecDone := FALSE;

                   #lastSeq := #KukaControlCmdSeq;          // <-- memoriza!
                   #lastCode := #code_int;             // memoriza qué comando es (para actualizar activos en DONE)

                   #state := 20;                    // BUSY
               END_IF; // bloqueo por pausa

               END_IF;

           END_IF;

       20: // BUSY

           #PlcStatusExecBusy := TRUE;

           IF ("rbDone" = "goTrigger") THEN
               // Fin confirmado por KUKA
               // 

               // Si venimos de CANCEL, este DONE es de cancelación
               IF #_cancelInFlight THEN
                   // comportamiento típico: marcar done "administrativo"
                   // (si prefieres diferenciar, añade PlcStatusExecCanceled)
                   #_cancelInFlight := FALSE;
               END_IF;

               #PlcStatusExecDone := TRUE;
               #PlcStatusExecBusy := FALSE;
               #PlcStatusExecAccepted := FALSE;
               // ACK de la orden completada
               #PlcStatusExecAckSeq := #lastSeq;

               // ✅ Actualiza activos al terminar de verdad
               //IF #lastCode = 201 THEN
                   //#PlcStatusActiveToolId := #toolReqId;
                //// ELSIF #lastCode = 202 THEN
                 ///  #PlcStatusActiveBaseId := #KukaControlCmdBaseRequestId;
              // ELSIF #lastCode = 203 THEN
                  // #PlcStatusActiveProfileId := #profileReqId;  // 
              // END_IF;

               // salir de pausa si termina un job por su curso natural
               #PlcStatusExecPaused := FALSE;

               #state := 0;                         // vuelve a IDLE

           END_IF;

       30: // DONE
           // limpiar y volver a IDLE
           #state := 0;


   END_CASE;
END_REGION
END_FUNCTION_BLOCK

// folder: 20. Robot Services/RobotPos

FUNCTION_BLOCK "TcpPoseDecoderLe32"   // FB4, LAD
{ S7_Optimized_Access := 'TRUE' }
VERSION : 0.1
// Decodifica con SWAP, convierte a DINT y escala.
   VAR_INPUT
      xIniRawLe : DWord;
      yIniRawLe : DWord;
      zIniRawLe : DWord;
      e1IniRawLe : DWord;
      xFinRawLe : DWord;
      yFinRawLe : DWord;
      zFinRawLe : DWord;
      e1FinRawLe : DWord;
      ToolActiveRawByte : Byte;
      BaseActiveRawByte : Byte;
   END_VAR
   VAR_OUTPUT
      tcpPosIniX_mm : LReal;
      tcpPosIniY_mm : LReal;
      tcpPosIniZ_mm : LReal;
      e1PosIni_mm : LReal;
      tcpPosFinX_mm : LReal;
      tcpPosFinY_mm : LReal;
      tcpPosFinZ_mm : LReal;
      e1PosFin_mm : LReal;
      toolActiveId : UDInt;
      baseActiveId : UDInt;
   END_VAR
   VAR_TEMP
      xIniDint : DInt;
      yIniDint : DInt;
      zIniDint : DInt;
      aDint : DInt;
      bDint : DInt;
      cDint : DInt;
      e1IniDint : DInt;
      xFinDint : DInt;
      yFinDint : DInt;
      zFinDint : DInt;
      e1FinDint : DInt;
   END_VAR
BEGIN

REGION Network 1 (SCL): // 1) Endianness: ABCD -> DCBA
   #xIniDint := DWORD_TO_DINT(SWAP(#xIniRawLe));
   #yIniDint := DWORD_TO_DINT(SWAP(#yIniRawLe));
   #zIniDint := DWORD_TO_DINT(SWAP(#zIniRawLe));

   #e1IniDint := DWORD_TO_DINT(SWAP(#e1IniRawLe));

   #xFinDint := DWORD_TO_DINT(SWAP(#xFinRawLe));
   #yFinDint := DWORD_TO_DINT(SWAP(#yFinRawLe));
   #zFinDint := DWORD_TO_DINT(SWAP(#zFinRawLe));
   #e1FinDint := DWORD_TO_DINT(SWAP(#e1FinRawLe));
END_REGION

REGION Network 2 (SCL): // 2) Escala fixed-point: µm->mm, mdeg->deg
   #tcpPosIniX_mm := DINT_TO_LREAL(#xIniDint) / 1000.0;
   #tcpPosIniY_mm := DINT_TO_LREAL(#yIniDint) / 1000.0;
   #tcpPosIniZ_mm := DINT_TO_LREAL(#zIniDint) / 1000.0;

   #e1PosIni_mm := DINT_TO_LREAL(#e1IniDint) / 1000.0;  // mm o deg según tu E1

